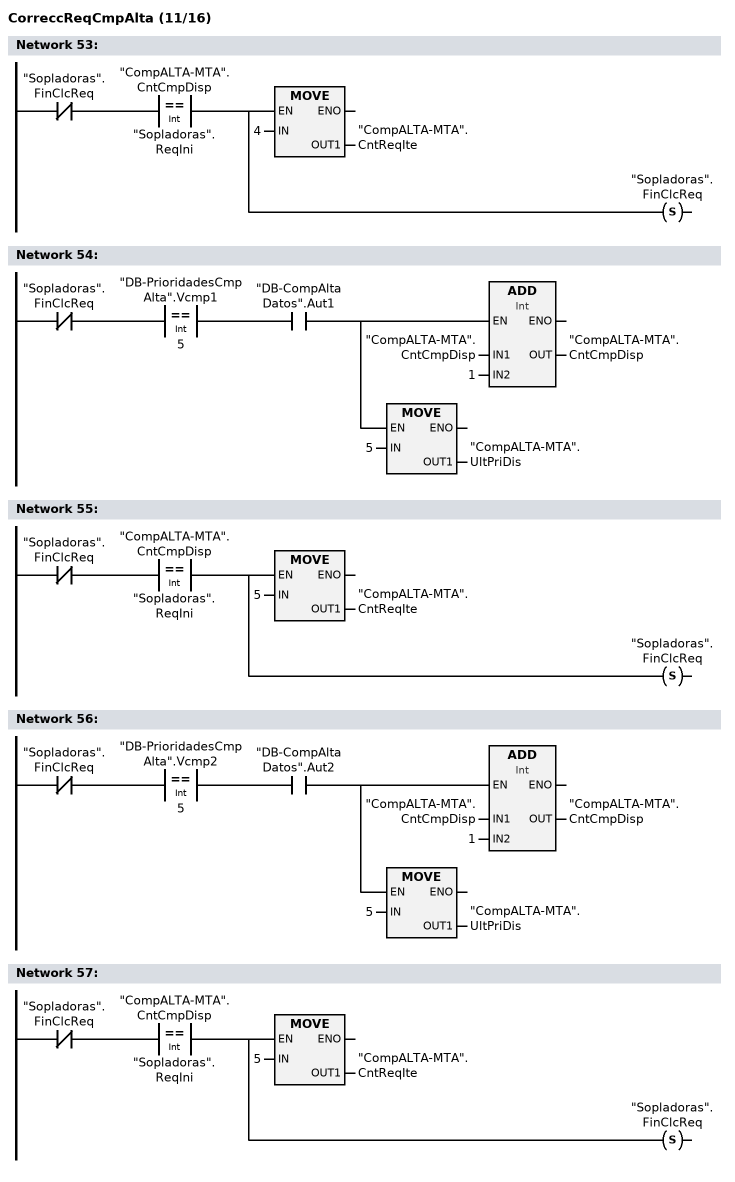
   RUNG wire#powerrail
      I_Contact( "Sopladoras".FinClcReq )
      { S7_Templates := "SrcType := Int" } EQ_Contact(in1 := "CompALTA-MTA".CntCmpDisp, in2 := "Sopladoras".ReqIni)
      wire#w1
      { S7_GenerateENO := "TRUE" } Move(in := 4, out1 => "CompALTA-MTA".CntReqIte)
   END_RUNG
   RUNG wire#w1
      S_Coil( "Sopladoras".FinClcReq )
   END_RUNG
   // the same network as SCL:
   IF NOT "Sopladoras".FinClcReq AND ("CompALTA-MTA".CntCmpDisp = "Sopladoras".ReqIni) THEN
       "CompALTA-MTA".CntReqIte := 4;
       "Sopladoras".FinClcReq := TRUE;
   END_IF;
END_REGION

REGION Network 54
   IF NOT "Sopladoras".FinClcReq AND ("DB-PrioridadesCmpAlta".Vcmp1 = 5) AND "DB-CompAltaDatos".Aut1 THEN
       "CompALTA-MTA".CntCmpDisp := "CompALTA-MTA".CntCmpDisp + 1;
       "CompALTA-MTA".UltPriDis := 5;
   END_IF;
END_REGION

REGION Network 55
   IF NOT "Sopladoras".FinClcReq AND ("CompALTA-MTA".CntCmpDisp = "Sopladoras".ReqIni) THEN
       "CompALTA-MTA".CntReqIte := 5;
       "Sopladoras".FinClcReq := TRUE;
   END_IF;
END_REGION

REGION Network 56
   IF NOT "Sopladoras".FinClcReq AND ("DB-PrioridadesCmpAlta".Vcmp2 = 5) AND "DB-CompAltaDatos".Aut2 THEN
       "CompALTA-MTA".CntCmpDisp := "CompALTA-MTA".CntCmpDisp + 1;
       "CompALTA-MTA".UltPriDis := 5;
   END_IF;
END_REGION

REGION Network 57
   IF NOT "Sopladoras".FinClcReq AND ("CompALTA-MTA".CntCmpDisp = "Sopladoras".ReqIni) THEN
       "CompALTA-MTA".CntReqIte := 5;
       "Sopladoras".FinClcReq := TRUE;
   END_IF;
END_REGION

REGION Network 58
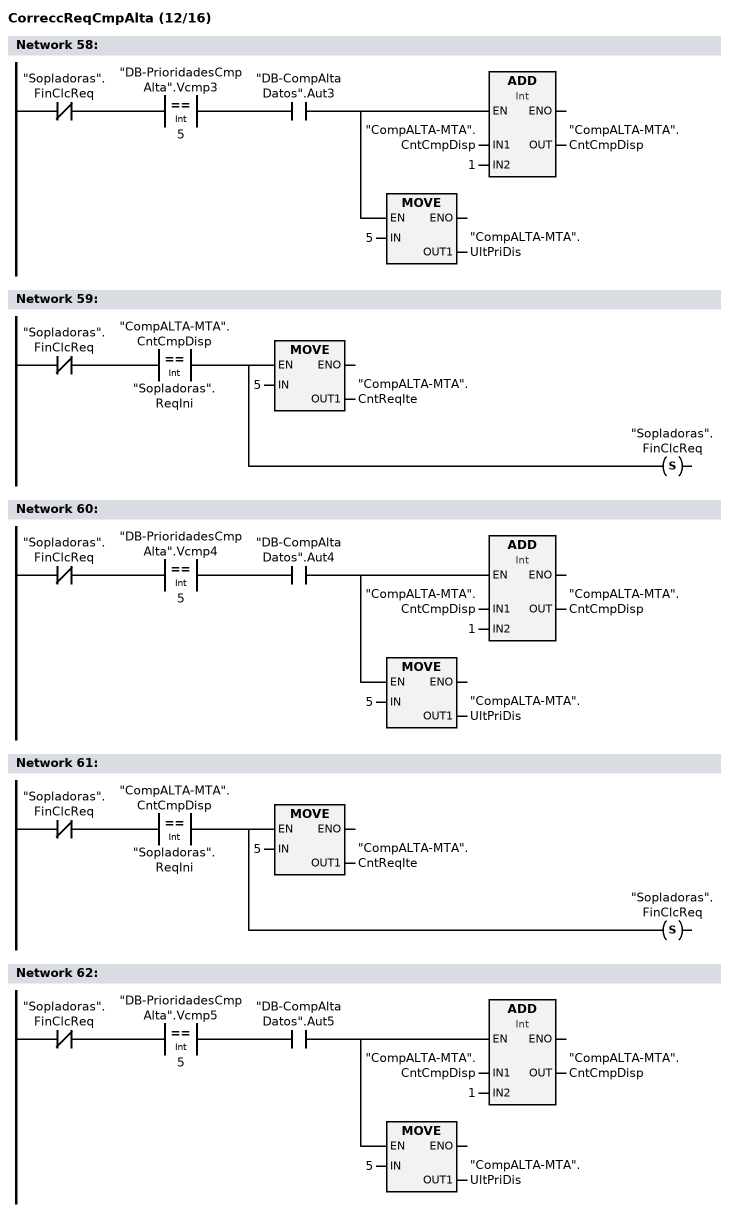
   IF NOT "Sopladoras".FinClcReq AND ("DB-PrioridadesCmpAlta".Vcmp3 = 5) AND "DB-CompAltaDatos".Aut3 THEN
       "CompALTA-MTA".CntCmpDisp := "CompALTA-MTA".CntCmpDisp + 1;
       "CompALTA-MTA".UltPriDis := 5;
   END_IF;
END_REGION

REGION Network 59
   IF NOT "Sopladoras".FinClcReq AND ("CompALTA-MTA".CntCmpDisp = "Sopladoras".ReqIni) THEN
       "CompALTA-MTA".CntReqIte := 5;
       "Sopladoras".FinClcReq := TRUE;
   END_IF;
END_REGION

REGION Network 60
   IF NOT "Sopladoras".FinClcReq AND ("DB-PrioridadesCmpAlta".Vcmp4 = 5) AND "DB-CompAltaDatos".Aut4 THEN
       "CompALTA-MTA".CntCmpDisp := "CompALTA-MTA".CntCmpDisp + 1;
       "CompALTA-MTA".UltPriDis := 5;
   END_IF;
END_REGION

REGION Network 61
   IF NOT "Sopladoras".FinClcReq AND ("CompALTA-MTA".CntCmpDisp = "Sopladoras".ReqIni) THEN
       "CompALTA-MTA".CntReqIte := 5;
       "Sopladoras".FinClcReq := TRUE;
   END_IF;
END_REGION

REGION Network 62
   IF NOT "Sopladoras".FinClcReq AND ("DB-PrioridadesCmpAlta".Vcmp5 = 5) AND "DB-CompAltaDatos".Aut5 THEN
       "CompALTA-MTA".CntCmpDisp := "CompALTA-MTA".CntCmpDisp + 1;
       "CompALTA-MTA".UltPriDis := 5;
   END_IF;
END_REGION

REGION Network 63
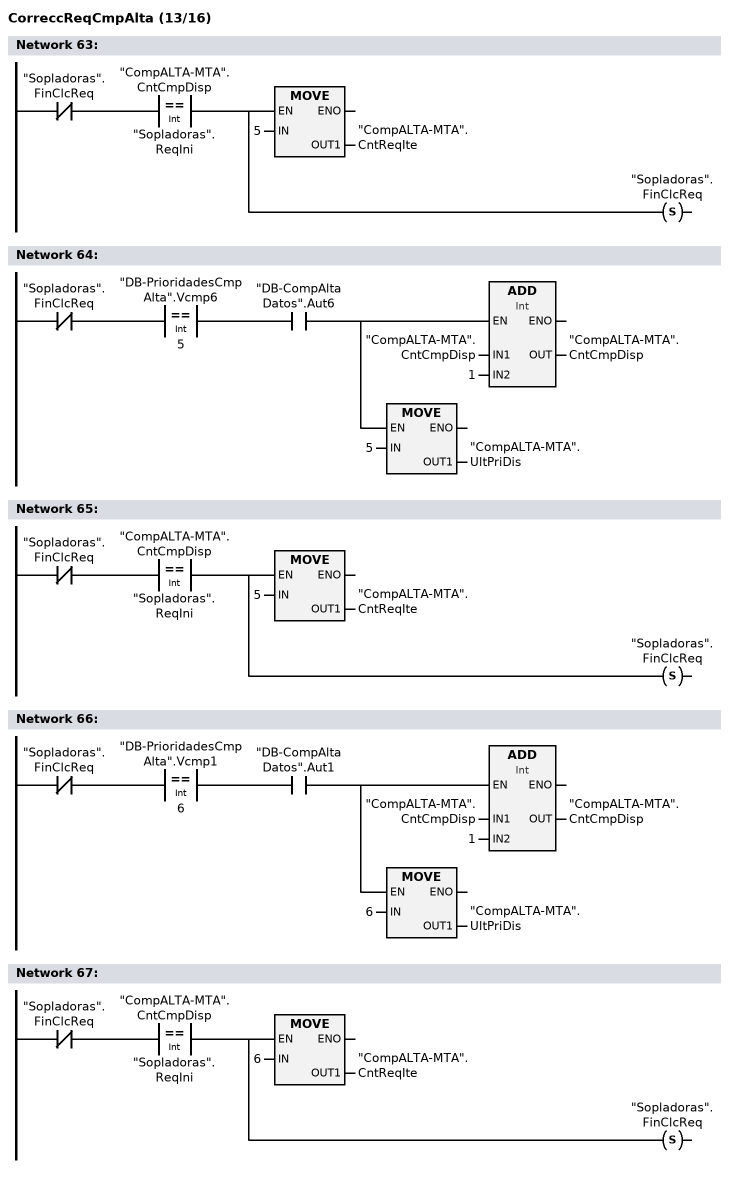
   IF NOT "Sopladoras".FinClcReq AND ("CompALTA-MTA".CntCmpDisp = "Sopladoras".ReqIni) THEN
       "CompALTA-MTA".CntReqIte := 5;
       "Sopladoras".FinClcReq := TRUE;
   END_IF;
END_REGION

REGION Network 64
   RUNG wire#powerrail
      I_Contact( "Sopladoras".FinClcReq )
      { S7_Templates := "SrcType := Int" } EQ_Contact(in1 := "DB-PrioridadesCmpAlta".Vcmp6, in2 := 5)
      Contact( "DB-CompAltaDatos".Aut6 )
      wire#w1
      { S7_Templates := "SrcType := Int"; S7_GenerateENO := "TRUE" } Add(in1 := "CompALTA-MTA".CntCmpDisp, in2 := 1, out => "CompALTA-MTA".CntCmpDisp)
   END_RUNG
   RUNG wire#w1
      { S7_GenerateENO := "TRUE" } Move(in := 5, out1 => "CompALTA-MTA".UltPriDis)
   END_RUNG
   // the same network as SCL:
   IF NOT "Sopladoras".FinClcReq AND ("DB-PrioridadesCmpAlta".Vcmp6 = 5) AND "DB-CompAltaDatos".Aut6 THEN
       "CompALTA-MTA".CntCmpDisp := "CompALTA-MTA".CntCmpDisp + 1;
       "CompALTA-MTA".UltPriDis := 5;
   END_IF;
END_REGION

REGION Network 65
   RUNG wire#powerrail
      I_Contact( "Sopladoras".FinClcReq )
      { S7_Templates := "SrcType := Int" } EQ_Contact(in1 := "CompALTA-MTA".CntCmpDisp, in2 := "Sopladoras".ReqIni)
      wire#w1
      { S7_GenerateENO := "TRUE" } Move(in := 5, out1 => "CompALTA-MTA".CntReqIte)
   END_RUNG
   RUNG wire#w1
      S_Coil( "Sopladoras".FinClcReq )
   END_RUNG
   // the same network as SCL:
   IF NOT "Sopladoras".FinClcReq AND ("CompALTA-MTA".CntCmpDisp = "Sopladoras".ReqIni) THEN
       "CompALTA-MTA".CntReqIte := 5;
       "Sopladoras".FinClcReq := TRUE;
   END_IF;
END_REGION

REGION Network 66
   RUNG wire#powerrail
      I_Contact( "Sopladoras".FinClcReq )
      { S7_Templates := "SrcType := Int" } EQ_Contact(in1 := "DB-PrioridadesCmpAlta".Vcmp1, in2 := 6)
      Contact( "DB-CompAltaDatos".Aut1 )
      wire#w1
      { S7_Templates := "SrcType := Int"; S7_GenerateENO := "TRUE" } Add(in1 := "CompALTA-MTA".CntCmpDisp, in2 := 1, out => "CompALTA-MTA".CntCmpDisp)
   END_RUNG
   RUNG wire#w1
      { S7_GenerateENO := "TRUE" } Move(in := 6, out1 => "CompALTA-MTA".UltPriDis)
   END_RUNG
   // the same network as SCL:
   IF NOT "Sopladoras".FinClcReq AND ("DB-PrioridadesCmpAlta".Vcmp1 = 6) AND "DB-CompAltaDatos".Aut1 THEN
       "CompALTA-MTA".CntCmpDisp := "CompALTA-MTA".CntCmpDisp + 1;
       "CompALTA-MTA".UltPriDis := 6;
   END_IF;
END_REGION

REGION Network 67
   RUNG wire#powerrail
      I_Contact( "Sopladoras".FinClcReq )
      { S7_Templates := "SrcType := Int" } EQ_Contact(in1 := "CompALTA-MTA".CntCmpDisp, in2 := "Sopladoras".ReqIni)
      wire#w1
      { S7_GenerateENO := "TRUE" } Move(in := 6, out1 => "CompALTA-MTA".CntReqIte)
   END_RUNG
   RUNG wire#w1
      S_Coil( "Sopladoras".FinClcReq )
   END_RUNG
   // the same network as SCL:
   IF NOT "Sopladoras".FinClcReq AND ("CompALTA-MTA".CntCmpDisp = "Sopladoras".ReqIni) THEN
       "CompALTA-MTA".CntReqIte := 6;
       "Sopladoras".FinClcReq := TRUE;
   END_IF;
END_REGION

REGION Network 68
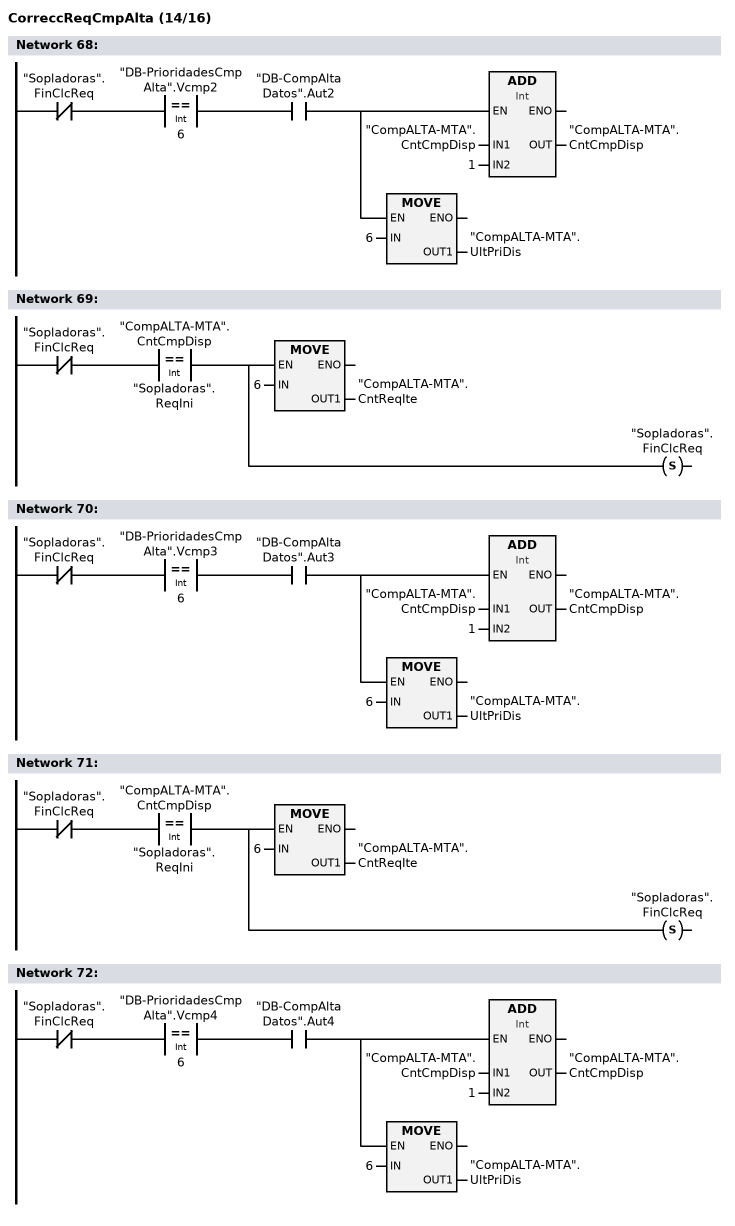
   RUNG wire#powerrail
      I_Contact( "Sopladoras".FinClcReq )
      { S7_Templates := "SrcType := Int" } EQ_Contact(in1 := "DB-PrioridadesCmpAlta".Vcmp2, in2 := 6)
      Contact( "DB-CompAltaDatos".Aut2 )
      wire#w1
      { S7_Templates := "SrcType := Int"; S7_GenerateENO := "TRUE" } Add(in1 := "CompALTA-MTA".CntCmpDisp, in2 := 1, out => "CompALTA-MTA".CntCmpDisp)
   END_RUNG
   RUNG wire#w1
      { S7_GenerateENO := "TRUE" } Move(in := 6, out1 => "CompALTA-MTA".UltPriDis)
   END_RUNG
   // the same network as SCL:
   IF NOT "Sopladoras".FinClcReq AND ("DB-PrioridadesCmpAlta".Vcmp2 = 6) AND "DB-CompAltaDatos".Aut2 THEN
       "CompALTA-MTA".CntCmpDisp := "CompALTA-MTA".CntCmpDisp + 1;
       "CompALTA-MTA".UltPriDis := 6;
   END_IF;
END_REGION

REGION Network 69
   RUNG wire#powerrail
      I_Contact( "Sopladoras".FinClcReq )
      { S7_Templates := "SrcType := Int" } EQ_Contact(in1 := "CompALTA-MTA".CntCmpDisp, in2 := "Sopladoras".ReqIni)
      wire#w1
      { S7_GenerateENO := "TRUE" } Move(in := 6, out1 => "CompALTA-MTA".CntReqIte)
   END_RUNG
   RUNG wire#w1
      S_Coil( "Sopladoras".FinClcReq )
   END_RUNG
   // the same network as SCL:
   IF NOT "Sopladoras".FinClcReq AND ("CompALTA-MTA".CntCmpDisp = "Sopladoras".ReqIni) THEN
       "CompALTA-MTA".CntReqIte := 6;
       "Sopladoras".FinClcReq := TRUE;
   END_IF;
END_REGION

REGION Network 70
   RUNG wire#powerrail
      I_Contact( "Sopladoras".FinClcReq )
      { S7_Templates := "SrcType := Int" } EQ_Contact(in1 := "DB-PrioridadesCmpAlta".Vcmp3, in2 := 6)
      Contact( "DB-CompAltaDatos".Aut3 )
      wire#w1
      { S7_Templates := "SrcType := Int"; S7_GenerateENO := "TRUE" } Add(in1 := "CompALTA-MTA".CntCmpDisp, in2 := 1, out => "CompALTA-MTA".CntCmpDisp)
   END_RUNG
   RUNG wire#w1
      { S7_GenerateENO := "TRUE" } Move(in := 6, out1 => "CompALTA-MTA".UltPriDis)
   END_RUNG
   // the same network as SCL:
   IF NOT "Sopladoras".FinClcReq AND ("DB-PrioridadesCmpAlta".Vcmp3 = 6) AND "DB-CompAltaDatos".Aut3 THEN
       "CompALTA-MTA".CntCmpDisp := "CompALTA-MTA".CntCmpDisp + 1;
       "CompALTA-MTA".UltPriDis := 6;
   END_IF;
END_REGION

REGION Network 71
   RUNG wire#powerrail
      I_Contact( "Sopladoras".FinClcReq )
      { S7_Templates := "SrcType := Int" } EQ_Contact(in1 := "CompALTA-MTA".CntCmpDisp, in2 := "Sopladoras".ReqIni)
      wire#w1
      { S7_GenerateENO := "TRUE" } Move(in := 6, out1 => "CompALTA-MTA".CntReqIte)
   END_RUNG
   RUNG wire#w1
      S_Coil( "Sopladoras".FinClcReq )
   END_RUNG
   // the same network as SCL:
   IF NOT "Sopladoras".FinClcReq AND ("CompALTA-MTA".CntCmpDisp = "Sopladoras".ReqIni) THEN
       "CompALTA-MTA".CntReqIte := 6;
       "Sopladoras".FinClcReq := TRUE;
   END_IF;
END_REGION

REGION Network 72
   RUNG wire#powerrail
      I_Contact( "Sopladoras".FinClcReq )
      { S7_Templates := "SrcType := Int" } EQ_Contact(in1 := "DB-PrioridadesCmpAlta".Vcmp4, in2 := 6)
      Contact( "DB-CompAltaDatos".Aut4 )
      wire#w1
      { S7_Templates := "SrcType := Int"; S7_GenerateENO := "TRUE" } Add(in1 := "CompALTA-MTA".CntCmpDisp, in2 := 1, out => "CompALTA-MTA".CntCmpDisp)
   END_RUNG
   RUNG wire#w1
      { S7_GenerateENO := "TRUE" } Move(in := 6, out1 => "CompALTA-MTA".UltPriDis)
   END_RUNG
   // the same network as SCL:
   IF NOT "Sopladoras".FinClcReq AND ("DB-PrioridadesCmpAlta".Vcmp4 = 6) AND "DB-CompAltaDatos".Aut4 THEN
       "CompALTA-MTA".CntCmpDisp := "CompALTA-MTA".CntCmpDisp + 1;
       "CompALTA-MTA".UltPriDis := 6;
   END_IF;
END_REGION

REGION Network 73
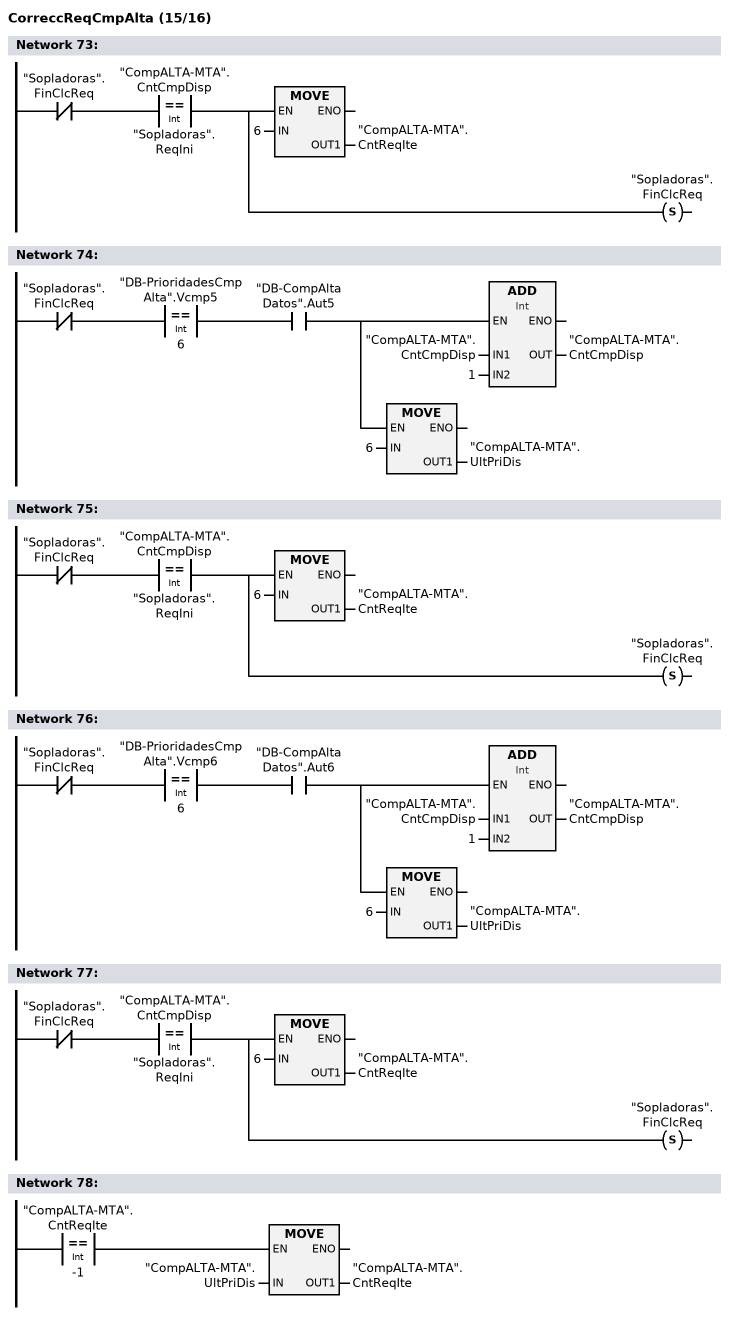
   RUNG wire#powerrail
      I_Contact( "Sopladoras".FinClcReq )
      { S7_Templates := "SrcType := Int" } EQ_Contact(in1 := "CompALTA-MTA".CntCmpDisp, in2 := "Sopladoras".ReqIni)
      wire#w1
      { S7_GenerateENO := "TRUE" } Move(in := 6, out1 => "CompALTA-MTA".CntReqIte)
   END_RUNG
   RUNG wire#w1
      S_Coil( "Sopladoras".FinClcReq )
   END_RUNG
   // the same network as SCL:
   IF NOT "Sopladoras".FinClcReq AND ("CompALTA-MTA".CntCmpDisp = "Sopladoras".ReqIni) THEN
       "CompALTA-MTA".CntReqIte := 6;
       "Sopladoras".FinClcReq := TRUE;
   END_IF;
END_REGION

REGION Network 74
   RUNG wire#powerrail
      I_Contact( "Sopladoras".FinClcReq )
      { S7_Templates := "SrcType := Int" } EQ_Contact(in1 := "DB-PrioridadesCmpAlta".Vcmp5, in2 := 6)
      Contact( "DB-CompAltaDatos".Aut5 )
      wire#w1
      { S7_Templates := "SrcType := Int"; S7_GenerateENO := "TRUE" } Add(in1 := "CompALTA-MTA".CntCmpDisp, in2 := 1, out => "CompALTA-MTA".CntCmpDisp)
   END_RUNG
   RUNG wire#w1
      { S7_GenerateENO := "TRUE" } Move(in := 6, out1 => "CompALTA-MTA".UltPriDis)
   END_RUNG
   // the same network as SCL:
   IF NOT "Sopladoras".FinClcReq AND ("DB-PrioridadesCmpAlta".Vcmp5 = 6) AND "DB-CompAltaDatos".Aut5 THEN
       "CompALTA-MTA".CntCmpDisp := "CompALTA-MTA".CntCmpDisp + 1;
       "CompALTA-MTA".UltPriDis := 6;
   END_IF;
END_REGION

REGION Network 75
   RUNG wire#powerrail
      I_Contact( "Sopladoras".FinClcReq )
      { S7_Templates := "SrcType := Int" } EQ_Contact(in1 := "CompALTA-MTA".CntCmpDisp, in2 := "Sopladoras".ReqIni)
      wire#w1
      { S7_GenerateENO := "TRUE" } Move(in := 6, out1 => "CompALTA-MTA".CntReqIte)
   END_RUNG
   RUNG wire#w1
      S_Coil( "Sopladoras".FinClcReq )
   END_RUNG
   // the same network as SCL:
   IF NOT "Sopladoras".FinClcReq AND ("CompALTA-MTA".CntCmpDisp = "Sopladoras".ReqIni) THEN
       "CompALTA-MTA".CntReqIte := 6;
       "Sopladoras".FinClcReq := TRUE;
   END_IF;
END_REGION

REGION Network 76
   RUNG wire#powerrail
      I_Contact( "Sopladoras".FinClcReq )
      { S7_Templates := "SrcType := Int" } EQ_Contact(in1 := "DB-PrioridadesCmpAlta".Vcmp6, in2 := 6)
      Contact( "DB-CompAltaDatos".Aut6 )
      wire#w1
      { S7_Templates := "SrcType := Int"; S7_GenerateENO := "TRUE" } Add(in1 := "CompALTA-MTA".CntCmpDisp, in2 := 1, out => "CompALTA-MTA".CntCmpDisp)
   END_RUNG
   RUNG wire#w1
      { S7_GenerateENO := "TRUE" } Move(in := 6, out1 => "CompALTA-MTA".UltPriDis)
   END_RUNG
   // the same network as SCL:
   IF NOT "Sopladoras".FinClcReq AND ("DB-PrioridadesCmpAlta".Vcmp6 = 6) AND "DB-CompAltaDatos".Aut6 THEN
       "CompALTA-MTA".CntCmpDisp := "CompALTA-MTA".CntCmpDisp + 1;
       "CompALTA-MTA".UltPriDis := 6;
   END_IF;
END_REGION

REGION Network 77
   RUNG wire#powerrail
      I_Contact( "Sopladoras".FinClcReq )
      { S7_Templates := "SrcType := Int" } EQ_Contact(in1 := "CompALTA-MTA".CntCmpDisp, in2 := "Sopladoras".ReqIni)
      wire#w1
      { S7_GenerateENO := "TRUE" } Move(in := 6, out1 => "CompALTA-MTA".CntReqIte)
   END_RUNG
   RUNG wire#w1
      S_Coil( "Sopladoras".FinClcReq )
   END_RUNG
   // the same network as SCL:
   IF NOT "Sopladoras".FinClcReq AND ("CompALTA-MTA".CntCmpDisp = "Sopladoras".ReqIni) THEN
       "CompALTA-MTA".CntReqIte := 6;
       "Sopladoras".FinClcReq := TRUE;
   END_IF;
END_REGION

REGION Network 78
   RUNG wire#powerrail
      { S7_Templates := "SrcType := Int" } EQ_Contact(in1 := "CompALTA-MTA".CntReqIte, in2 := -1)
      { S7_GenerateENO := "TRUE" } Move(in := "CompALTA-MTA".UltPriDis, out1 => "CompALTA-MTA".CntReqIte)
   END_RUNG
   // the same network as SCL:
   IF "CompALTA-MTA".CntReqIte = (-1) THEN "CompALTA-MTA".CntReqIte := "CompALTA-MTA".UltPriDis; END_IF;
END_REGION

REGION Network 79
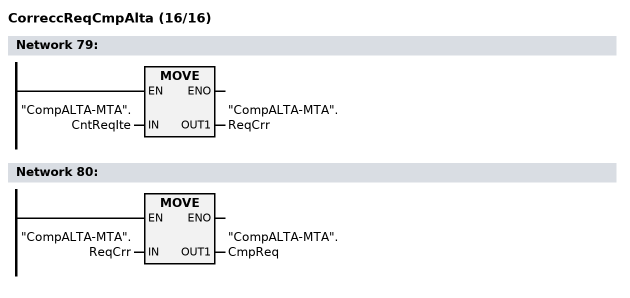
   RUNG wire#powerrail
      { S7_GenerateENO := "TRUE" } Move(in := "CompALTA-MTA".CntReqIte, out1 => "CompALTA-MTA".ReqCrr)
   END_RUNG
   // the same network as SCL:
   "CompALTA-MTA".ReqCrr := "CompALTA-MTA".CntReqIte;
END_REGION

REGION Network 80
   RUNG wire#powerrail
      { S7_GenerateENO := "TRUE" } Move(in := "CompALTA-MTA".ReqCrr, out1 => "CompALTA-MTA".CmpReq)
   END_RUNG
   // the same network as SCL:
   "CompALTA-MTA".CmpReq := "CompALTA-MTA".ReqCrr;
END_REGION
END_FUNCTION

FUNCTION "CalcEst6" : Void   // FC50, LAD
{ S7_Optimized_Access := 'FALSE' }
VERSION : 0.1
   VAR_TEMP   // added for the SCL form of the ladder/FBD networks
      _w1 : Bool;
   END_VAR
BEGIN

REGION Network 1: Prioritaria 1
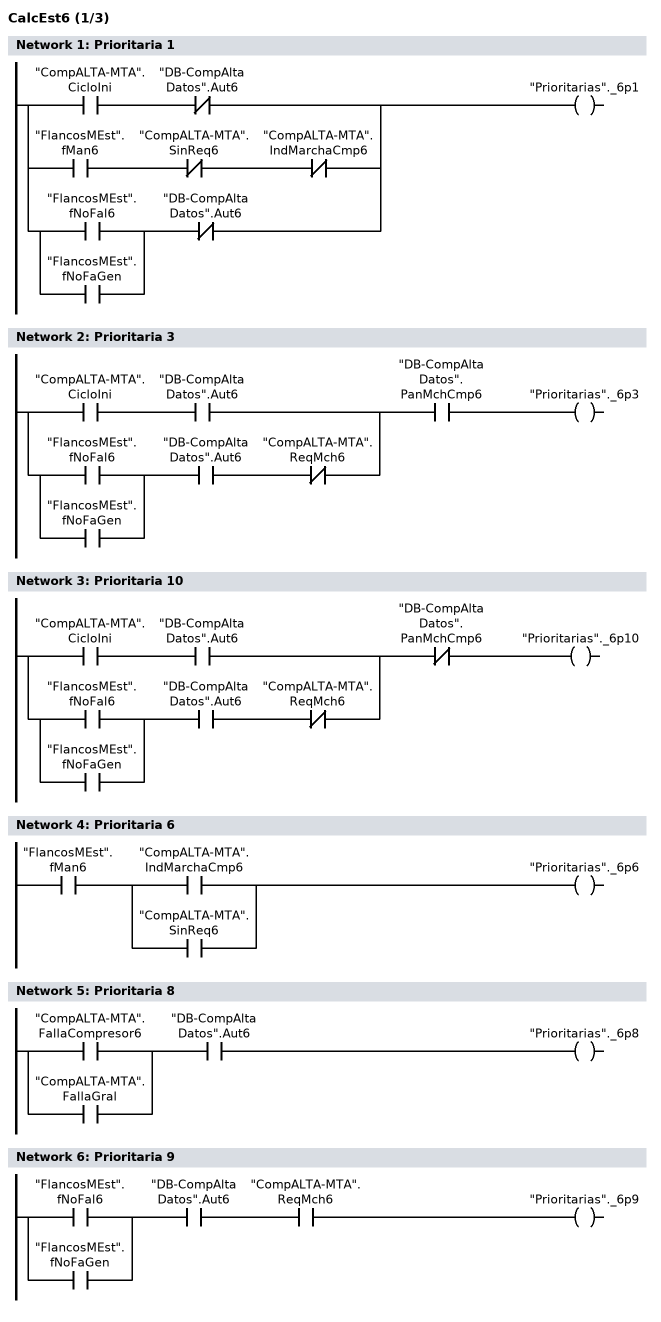
   RUNG wire#powerrail
      Contact( "CompALTA-MTA".CicloIni )
      I_Contact( "DB-CompAltaDatos".Aut6 )
      wire#w1
      Coil( "Prioritarias"._6p1 )
   END_RUNG
   RUNG wire#powerrail
      Contact( "FlancosMEst".fMan6 )
      I_Contact( "CompALTA-MTA".SinReq6 )
      I_Contact( "CompALTA-MTA".IndMarchaCmp6 )
   END_RUNG wire#w1
   RUNG wire#powerrail
      Contact( "FlancosMEst".fNoFal6 )
      wire#w2
      I_Contact( "DB-CompAltaDatos".Aut6 )
   END_RUNG wire#w1
   RUNG wire#powerrail
      Contact( "FlancosMEst".fNoFaGen )
   END_RUNG wire#w2
   // the same network as SCL:
   "Prioritarias"._6p1 := ("CompALTA-MTA".CicloIni AND NOT "DB-CompAltaDatos".Aut6) OR ("FlancosMEst".fMan6 AND NOT "CompALTA-MTA".SinReq6 AND NOT "CompALTA-MTA".IndMarchaCmp6) OR (("FlancosMEst".fNoFal6 OR "FlancosMEst".fNoFaGen) AND NOT "DB-CompAltaDatos".Aut6);
END_REGION

REGION Network 2: Prioritaria 3
   RUNG wire#powerrail
      Contact( "CompALTA-MTA".CicloIni )
      Contact( "DB-CompAltaDatos".Aut6 )
      wire#w1
      Contact( "DB-CompAltaDatos".PanMchCmp6 )
      Coil( "Prioritarias"._6p3 )
   END_RUNG
   RUNG wire#powerrail
      Contact( "FlancosMEst".fNoFal6 )
      wire#w2
      Contact( "DB-CompAltaDatos".Aut6 )
      I_Contact( "CompALTA-MTA".ReqMch6 )
   END_RUNG wire#w1
   RUNG wire#powerrail
      Contact( "FlancosMEst".fNoFaGen )
   END_RUNG wire#w2
   // the same network as SCL:
   "Prioritarias"._6p3 := (("CompALTA-MTA".CicloIni AND "DB-CompAltaDatos".Aut6) OR (("FlancosMEst".fNoFal6 OR "FlancosMEst".fNoFaGen) AND "DB-CompAltaDatos".Aut6 AND NOT "CompALTA-MTA".ReqMch6)) AND "DB-CompAltaDatos".PanMchCmp6;
END_REGION

REGION Network 3: Prioritaria 10
   RUNG wire#powerrail
      Contact( "CompALTA-MTA".CicloIni )
      Contact( "DB-CompAltaDatos".Aut6 )
      wire#w1
      I_Contact( "DB-CompAltaDatos".PanMchCmp6 )
      Coil( "Prioritarias"._6p10 )
   END_RUNG
   RUNG wire#powerrail
      Contact( "FlancosMEst".fNoFal6 )
      wire#w2
      Contact( "DB-CompAltaDatos".Aut6 )
      I_Contact( "CompALTA-MTA".ReqMch6 )
   END_RUNG wire#w1
   RUNG wire#powerrail
      Contact( "FlancosMEst".fNoFaGen )
   END_RUNG wire#w2
   // the same network as SCL:
   "Prioritarias"._6p10 := (("CompALTA-MTA".CicloIni AND "DB-CompAltaDatos".Aut6) OR (("FlancosMEst".fNoFal6 OR "FlancosMEst".fNoFaGen) AND "DB-CompAltaDatos".Aut6 AND NOT "CompALTA-MTA".ReqMch6)) AND NOT "DB-CompAltaDatos".PanMchCmp6;
END_REGION

REGION Network 4: Prioritaria 6
   RUNG wire#powerrail
      Contact( "FlancosMEst".fMan6 )
      wire#w1
      Contact( "CompALTA-MTA".IndMarchaCmp6 )
      wire#w2
      Coil( "Prioritarias"._6p6 )
   END_RUNG
   RUNG wire#w1
      Contact( "CompALTA-MTA".SinReq6 )
   END_RUNG wire#w2
   // the same network as SCL:
   "Prioritarias"._6p6 := "FlancosMEst".fMan6 AND ("CompALTA-MTA".IndMarchaCmp6 OR "CompALTA-MTA".SinReq6);
END_REGION

REGION Network 5: Prioritaria 8
   RUNG wire#powerrail
      Contact( "CompALTA-MTA".FallaCompresor6 )
      wire#w1
      Contact( "DB-CompAltaDatos".Aut6 )
      Coil( "Prioritarias"._6p8 )
   END_RUNG
   RUNG wire#powerrail
      Contact( "CompALTA-MTA".FallaGral )
   END_RUNG wire#w1
   // the same network as SCL:
   "Prioritarias"._6p8 := ("CompALTA-MTA".FallaCompresor6 OR "CompALTA-MTA".FallaGral) AND "DB-CompAltaDatos".Aut6;
END_REGION

REGION Network 6: Prioritaria 9
   RUNG wire#powerrail
      Contact( "FlancosMEst".fNoFal6 )
      wire#w1
      Contact( "DB-CompAltaDatos".Aut6 )
      Contact( "CompALTA-MTA".ReqMch6 )
      Coil( "Prioritarias"._6p9 )
   END_RUNG
   RUNG wire#powerrail
      Contact( "FlancosMEst".fNoFaGen )
   END_RUNG wire#w1
   // the same network as SCL:
   "Prioritarias"._6p9 := ("FlancosMEst".fNoFal6 OR "FlancosMEst".fNoFaGen) AND "DB-CompAltaDatos".Aut6 AND "CompALTA-MTA".ReqMch6;
END_REGION

REGION Network 7: Concatenadora 1
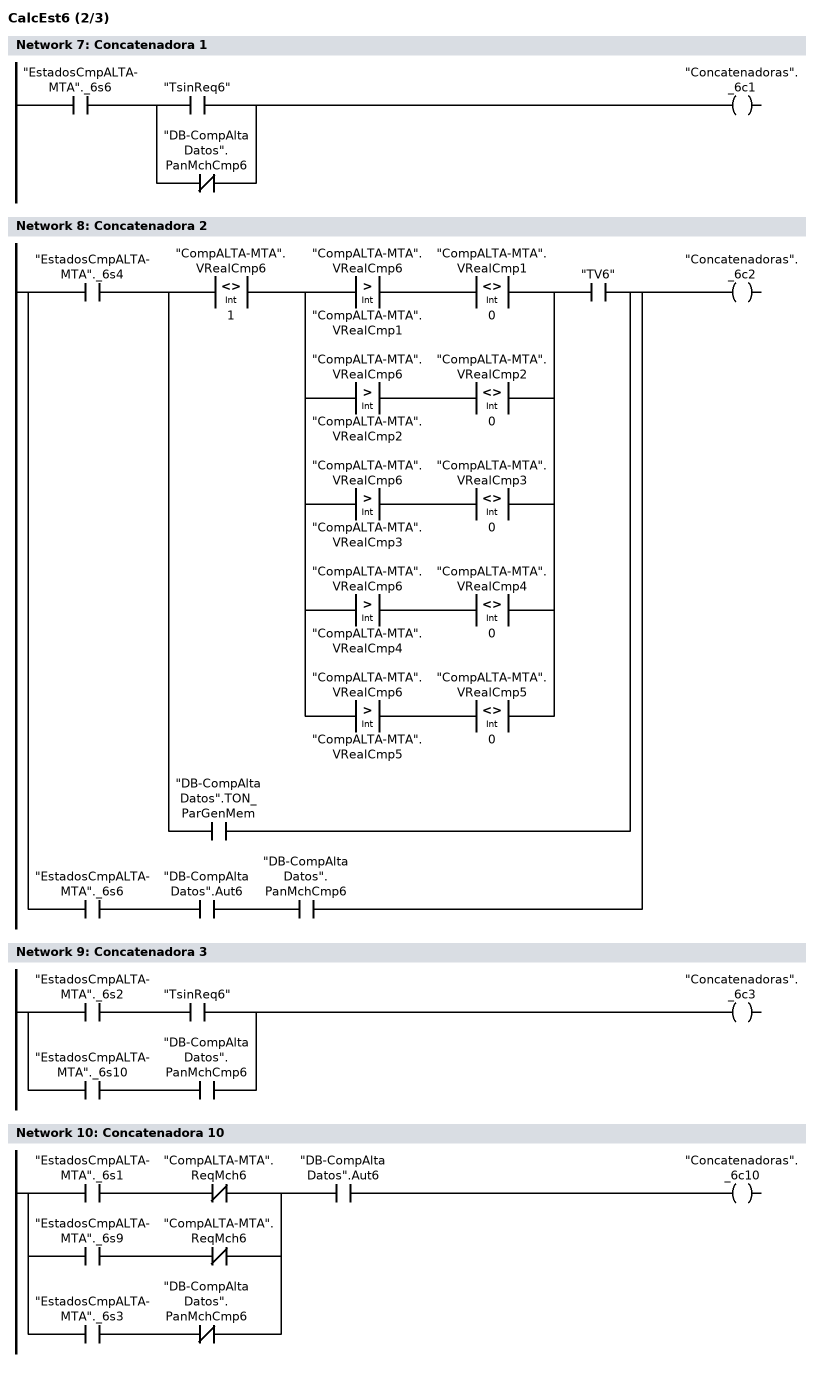
   RUNG wire#powerrail
      Contact( "EstadosCmpALTA-MTA"._6s6 )
      wire#w1
      Contact( "TsinReq6" )
      wire#w2
      Coil( "Concatenadoras"._6c1 )
   END_RUNG
   RUNG wire#w1
      I_Contact( "DB-CompAltaDatos".PanMchCmp6 )
   END_RUNG wire#w2
   // the same network as SCL:
   "Concatenadoras"._6c1 := "EstadosCmpALTA-MTA"._6s6 AND ("TsinReq6" OR NOT "DB-CompAltaDatos".PanMchCmp6);
END_REGION

REGION Network 8: Concatenadora 2
   RUNG wire#powerrail
      Contact( "EstadosCmpALTA-MTA"._6s4 )
      wire#w1
      { S7_Templates := "SrcType := Int" } NE_Contact(in1 := "CompALTA-MTA".VRealCmp6, in2 := 1)
      wire#w2
      { S7_Templates := "SrcType := Int" } GT_Contact(in1 := "CompALTA-MTA".VRealCmp6, in2 := "CompALTA-MTA".VRealCmp1)
      { S7_Templates := "SrcType := Int" } NE_Contact(in1 := "CompALTA-MTA".VRealCmp1, in2 := 0)
      wire#w3
      Contact( "TV6" )
      wire#w4
      Coil( "Concatenadoras"._6c2 )
   END_RUNG
   RUNG wire#w2
      { S7_Templates := "SrcType := Int" } GT_Contact(in1 := "CompALTA-MTA".VRealCmp6, in2 := "CompALTA-MTA".VRealCmp2)
      { S7_Templates := "SrcType := Int" } NE_Contact(in1 := "CompALTA-MTA".VRealCmp2, in2 := 0)
   END_RUNG wire#w3
   RUNG wire#w2
      { S7_Templates := "SrcType := Int" } GT_Contact(in1 := "CompALTA-MTA".VRealCmp6, in2 := "CompALTA-MTA".VRealCmp3)
      { S7_Templates := "SrcType := Int" } NE_Contact(in1 := "CompALTA-MTA".VRealCmp3, in2 := 0)
   END_RUNG wire#w3
   RUNG wire#w2
      { S7_Templates := "SrcType := Int" } GT_Contact(in1 := "CompALTA-MTA".VRealCmp6, in2 := "CompALTA-MTA".VRealCmp4)
      { S7_Templates := "SrcType := Int" } NE_Contact(in1 := "CompALTA-MTA".VRealCmp4, in2 := 0)
   END_RUNG wire#w3
   RUNG wire#w2
      { S7_Templates := "SrcType := Int" } GT_Contact(in1 := "CompALTA-MTA".VRealCmp6, in2 := "CompALTA-MTA".VRealCmp5)
      { S7_Templates := "SrcType := Int" } NE_Contact(in1 := "CompALTA-MTA".VRealCmp5, in2 := 0)
   END_RUNG wire#w3
   RUNG wire#w1
      Contact( "DB-CompAltaDatos".TON_ParGenMem )
   END_RUNG wire#w4
   RUNG wire#powerrail
      Contact( "EstadosCmpALTA-MTA"._6s6 )
      Contact( "DB-CompAltaDatos".Aut6 )
      Contact( "DB-CompAltaDatos".PanMchCmp6 )
   END_RUNG wire#w4
   // the same network as SCL:
   "Concatenadoras"._6c2 := ("EstadosCmpALTA-MTA"._6s4 AND ((("CompALTA-MTA".VRealCmp6 <> 1) AND ((("CompALTA-MTA".VRealCmp6 > "CompALTA-MTA".VRealCmp1) AND ("CompALTA-MTA".VRealCmp1 <> 0)) OR (("CompALTA-MTA".VRealCmp6 > "CompALTA-MTA".VRealCmp2) AND ("CompALTA-MTA".VRealCmp2 <> 0)) OR (("CompALTA-MTA".VRealCmp6 > "CompALTA-MTA".VRealCmp3) AND ("CompALTA-MTA".VRealCmp3 <> 0)) OR (("CompALTA-MTA".VRealCmp6 > "CompALTA-MTA".VRealCmp4) AND ("CompALTA-MTA".VRealCmp4 <> 0)) OR (("CompALTA-MTA".VRealCmp6 > "CompALTA-MTA".VRealCmp5) AND ("CompALTA-MTA".VRealCmp5 <> 0))) AND "TV6") OR "DB-CompAltaDatos".TON_ParGenMem)) OR ("EstadosCmpALTA-MTA"._6s6 AND "DB-CompAltaDatos".Aut6 AND "DB-CompAltaDatos".PanMchCmp6);
END_REGION

REGION Network 9: Concatenadora 3
   RUNG wire#powerrail
      Contact( "EstadosCmpALTA-MTA"._6s2 )
      Contact( "TsinReq6" )
      wire#w1
      Coil( "Concatenadoras"._6c3 )
   END_RUNG
   RUNG wire#powerrail
      Contact( "EstadosCmpALTA-MTA"._6s10 )
      Contact( "DB-CompAltaDatos".PanMchCmp6 )
   END_RUNG wire#w1
   // the same network as SCL:
   "Concatenadoras"._6c3 := ("EstadosCmpALTA-MTA"._6s2 AND "TsinReq6") OR ("EstadosCmpALTA-MTA"._6s10 AND "DB-CompAltaDatos".PanMchCmp6);
END_REGION
